      on Press: SetTag("MH_Control_Visibility", 1); SetTag("Press_Control_Screen", 2)
      Visibility <- "DB704_MH_Value_Mixinghead{0}_AmountComponent"
   Button "Button_31" at 489,499 size 94x25; TextOff 'Text'
      on Press: SetTag("MH_Control_Visibility", 2); SetTag("Temp_Control_Screen", 2)
      Visibility <- "DB704_MH_Value_Mixinghead{0}_AmountComponent"
   Button "Button_33" at 489,554 size 94x25; TextOff 'Text'
      on Press: SetTag("MH_Control_Visibility", 2); SetTag("Temp_Control_Screen", 4)
      Visibility <- "DB704_MH_Value_Mixinghead{0}_AmountComponent"
   Button "Button_32" at 489,527 size 94x25; TextOff 'bar'
      on Press: SetTag("MH_Control_Visibility", 1); SetTag("Press_Control_Screen", 4)
      Visibility <- "DB704_MH_Value_Mixinghead{0}_AmountComponent"
   Button "Button_6" at 768,446 size 94x25; TextOff 'Text'
      on Press: SetTag("MH_Control_Visibility", 2); SetTag("Temp_Control_Screen", 1)
      Visibility <- "DB704_MH_Value_Mixinghead{0}_AmountComponent"
   Button "Button_37" at 768,554 size 94x25; TextOff 'Text'
      on Press: SetTag("MH_Control_Visibility", 2); SetTag("Temp_Control_Screen", 5)
      Visibility <- "DB704_MH_Value_Mixinghead{0}_AmountComponent"
   Button "Button_36" at 768,527 size 94x25; TextOff 'bar'
      on Press: SetTag("MH_Control_Visibility", 1); SetTag("Press_Control_Screen", 5)
      Visibility <- "DB704_MH_Value_Mixinghead{0}_AmountComponent"
   Button "Button_35" at 768,499 size 94x25; TextOff 'Text'
      on Press: SetTag("MH_Control_Visibility", 2); SetTag("Temp_Control_Screen", 3)
      Visibility <- "DB704_MH_Value_Mixinghead{0}_AmountComponent"
   Button "Button_34" at 768,473 size 94x25; TextOff 'bar'
      on Press: SetTag("MH_Control_Visibility", 1); SetTag("Press_Control_Screen", 3)
      Visibility <- "DB704_MH_Value_Mixinghead{0}_AmountComponent"
   Button "Button_5" at 768,421 size 94x25; TextOff 'bar'
      on Press: SetTag("MH_Control_Visibility", 1); SetTag("Press_Control_Screen", 1)
      Visibility <- "DB704_MH_Value_Mixinghead{0}_AmountComponent"
   Button "Button_19" at 332,596 size 138x30; TextOff 'Text'; TextList "Pump_Name"
      Visibility <- "DB704_MH_Value_Mixinghead{0}_AmountComponent"
      ProcessValue <- "DB704_MH_Value_Mixinghead{0}_MH_Connection{1}_Pump_No"
      Appearance <- "DB614_MH_State_MH_Connection{0}_colour{1}"
   Button "Button_38" at 470,596 size 138x30; TextOff 'Text'; TextList "Pump_Name"
      Visibility <- "DB704_MH_Value_Mixinghead{0}_AmountComponent"
      ProcessValue <- "DB704_MH_Value_Mixinghead{0}_MH_Connection{2}_Pump_No"
      Appearance <- "DB614_MH_State_MH_Connection{0}_colour{2}"
   Button "Button_40" at 608,596 size 138x30; TextOff 'Text'; TextList "Pump_Name"
      Visibility <- "DB704_MH_Value_Mixinghead{0}_AmountComponent"
      ProcessValue <- "DB704_MH_Value_Mixinghead{0}_MH_Connection{3}_Pump_No"
      Appearance <- "DB614_MH_State_MH_Connection{0}_colour{3}"
   Button "Button_47" at 746,596 size 138x30; TextOff 'Text'; TextList "Pump_Name"
      Visibility <- "DB704_MH_Value_Mixinghead{0}_AmountComponent"
      ProcessValue <- "DB704_MH_Value_Mixinghead{0}_MH_Connection{4}_Pump_No"
      Appearance <- "DB614_MH_State_MH_Connection{0}_colour{4}"
   Button "Button_48" at 884,596 size 138x30; TextOff 'Text'; TextList "Pump_Name"
      Visibility <- "DB704_MH_Value_Mixinghead{0}_AmountComponent"
      ProcessValue <- "DB704_MH_Value_Mixinghead{0}_MH_Connection{5}_Pump_No"
      Appearance <- "DB614_MH_State_MH_Connection{0}_colour{5}"
   Button "Button_49" at 1022,596 size 138x30; TextOff 'Text'; TextList "Pump_Name"
      Visibility <- "DB704_MH_Value_Mixinghead{0}_AmountComponent"
      ProcessValue <- "DB704_MH_Value_Mixinghead{0}_MH_Connection{6}_Pump_No"
      Appearance <- "DB614_MH_State_MH_Connection{0}_colour{6}"
   Button "Button_50" at 342,413 size 138x30; TextOff 'Text'; TextList "Pump_Name"
      Visibility <- "DB704_MH_Value_Mixinghead{0}_AmountComponent"
      ProcessValue <- "DB704_MH_Value_Mixinghead{0}_MH_Connection{1}_Pump_No"
      Appearance <- "DB614_MH_State_MH_Connection{0}_colour{1}"
   Button "Button_51" at 342,474 size 138x30; TextOff 'Text'; TextList "Pump_Name"
      Visibility <- "DB704_MH_Value_Mixinghead{0}_AmountComponent"
      ProcessValue <- "DB704_MH_Value_Mixinghead{0}_MH_Connection{3}_Pump_No"
      Appearance <- "DB614_MH_State_MH_Connection{0}_colour{3}"
   Button "Button_52" at 342,535 size 138x30; TextOff 'Text'; TextList "Pump_Name"
      Visibility <- "DB704_MH_Value_Mixinghead{0}_AmountComponent"
      ProcessValue <- "DB704_MH_Value_Mixinghead{0}_MH_Connection{5}_Pump_No"
      Appearance <- "DB614_MH_State_MH_Connection{0}_colour{5}"
   Button "Button_53" at 871,413 size 138x30; TextOff 'Text'; TextList "Pump_Name"
      Visibility <- "DB704_MH_Value_Mixinghead{0}_AmountComponent"
      ProcessValue <- "DB704_MH_Value_Mixinghead{0}_MH_Connection{2}_Pump_No"
      Appearance <- "DB614_MH_State_MH_Connection{0}_colour{2}"
   Button "Button_54" at 871,474 size 138x30; TextOff 'Text'; TextList "Pump_Name"
      Visibility <- "DB704_MH_Value_Mixinghead{0}_AmountComponent"
      ProcessValue <- "DB704_MH_Value_Mixinghead{0}_MH_Connection{4}_Pump_No"
      Appearance <- "DB614_MH_State_MH_Connection{0}_colour{4}"
   Button "Button_55" at 871,535 size 138x30; TextOff 'Text'; TextList "Pump_Name"
      Visibility <- "DB704_MH_Value_Mixinghead{0}_AmountComponent"
      ProcessValue <- "DB704_MH_Value_Mixinghead{0}_MH_Connection{6}_Pump_No"
      Appearance <- "DB614_MH_State_MH_Connection{0}_colour{6}"
   GraphicView "Graphic view_10" at 600,423 size 40x37; Picture "logoff"
      Visibility <- "DB123_MH_IO_Signals_MH{0}_IN_MH_Prog_No_MH"
   TextField "Text field_54" at 838,273 size 46x25; Text 's'
      Visibility <- "DB704_MH_Value_Mixinghead{0}_Cleaning_Piston_CP_withInterval"
   TextField "Text field_55" at 838,303 size 46x25; Text 's'
      Visibility <- "DB704_MH_Value_Mixinghead{0}_Cleaning_Piston_CP_withInterval"
   TextField "Text field_40" at 202,455 size 94x25; Text 'NL'
      Visibility <- "DB704_MH_Value_Mixinghead{0}_WithInerting"
   TextField "Text field_41" at 202,430 size 94x25; Text 'NL'
      Visibility <- "DB704_MH_Value_Mixinghead{0}_WithInerting"
   Rectangle "Rectangle_11" at 332,627 size 138x40
      Visibility <- "DB614_MH_State_MH_Status{0}_QPB_Values_selected"
   Rectangle "Rectangle_12" at 332,666 size 138x40
      Visibility <- "DB614_MH_State_MH_Status{0}_QPB_Values_selected"
   Rectangle "Rectangle_13" at 332,705 size 138x40
      Visibility <- "DB614_MH_State_MH_Status{0}_QPB_Values_selected"
   Rectangle "Rectangle_14" at 332,744 size 138x40
      Visibility <- "DB614_MH_State_MH_Status{0}_QPB_Values_selected"
   Rectangle "Rectangle_7" at 470,627 size 138x40
      Visibility <- "DB614_MH_State_MH_Status{0}_QPB_Values_selected"
   Rectangle "Rectangle_8" at 470,666 size 138x40
      Visibility <- "DB614_MH_State_MH_Status{0}_QPB_Values_selected"
   Rectangle "Rectangle_9" at 470,705 size 138x40
      Visibility <- "DB614_MH_State_MH_Status{0}_QPB_Values_selected"
   Rectangle "Rectangle_10" at 470,744 size 138x40
      Visibility <- "DB614_MH_State_MH_Status{0}_QPB_Values_selected"
   TextField "Text field_10" at 106,635 size 70x25; Text 'actual:'
   TextField "Text field_11" at 106,673 size 93x25; Text 'Reduced:'
      Visibility <- "DB614_MH_State_MH_Status{0}_QPB_Values_selected"
   TextField "Text field_12" at 106,711 size 144x25; Text 'High pressure:'
      Visibility <- "DB614_MH_State_MH_Status{0}_QPB_Values_selected"
   TextField "Text field_13" at 106,752 size 139x25; Text 'Low pressure:'
      Visibility <- "DB614_MH_State_MH_Status{0}_QPB_Values_selected"
   TextField "Text field_14" at 277,635 size 46x25; Text 'g/s'
   TextField "Text field_16" at 277,673 size 46x25; Text 'g/s'
      Visibility <- "DB614_MH_State_MH_Status{0}_QPB_Values_selected"
   TextField "Text field_17" at 277,711 size 46x25; Text 'g/s'
      Visibility <- "DB614_MH_State_MH_Status{0}_QPB_Values_selected"
   TextField "Text field_18" at 277,749 size 46x25; Text 'bar'
      Visibility <- "DB614_MH_State_MH_Status{0}_QPB_Values_selected"
   Button "reduced icon" at 237,673 size 34x27; TextOff 'Text'; PictureOff "Reduced green"
      Visibility <- "DB614_MH_State_MH_Status{0}_QPB_Values_selected"
   Button "Interval icon" at 237,712 size 34x27; TextOff 'Text'; PictureOff "Interval green"
      Visibility <- "DB614_MH_State_MH_Status{0}_QPB_Values_selected"
   Button "Lowpress icon" at 237,751 size 34x27; TextOff 'Text'; PictureOff "Lowpress green"
      Visibility <- "DB614_MH_State_MH_Status{0}_QPB_Values_selected"
   Rectangle "Rectangle_15" at 608,627 size 138x40
      Visibility <- "DB614_MH_State_MH_Status{0}_QPB_Values_selected"
   Rectangle "Rectangle_16" at 608,666 size 138x40
      Visibility <- "DB614_MH_State_MH_Status{0}_QPB_Values_selected"
   Rectangle "Rectangle_17" at 608,705 size 138x40
      Visibility <- "DB614_MH_State_MH_Status{0}_QPB_Values_selected"
   Rectangle "Rectangle_18" at 608,744 size 138x40
      Visibility <- "DB614_MH_State_MH_Status{0}_QPB_Values_selected"
   Rectangle "Rectangle_19" at 746,627 size 138x40
      Visibility <- "DB614_MH_State_MH_Status{0}_QPB_Values_selected"
   Rectangle "Rectangle_20" at 746,666 size 138x40
      Visibility <- "DB614_MH_State_MH_Status{0}_QPB_Values_selected"
   Rectangle "Rectangle_21" at 746,705 size 138x40
      Visibility <- "DB614_MH_State_MH_Status{0}_QPB_Values_selected"
   Rectangle "Rectangle_22" at 746,744 size 138x40
      Visibility <- "DB614_MH_State_MH_Status{0}_QPB_Values_selected"
   Rectangle "Rectangle_23" at 884,627 size 138x40
      Visibility <- "DB614_MH_State_MH_Status{0}_QPB_Values_selected"
   Rectangle "Rectangle_24" at 884,666 size 138x40
      Visibility <- "DB614_MH_State_MH_Status{0}_QPB_Values_selected"
   Rectangle "Rectangle_25" at 884,705 size 138x40
      Visibility <- "DB614_MH_State_MH_Status{0}_QPB_Values_selected"
   Rectangle "Rectangle_26" at 884,744 size 138x40
      Visibility <- "DB614_MH_State_MH_Status{0}_QPB_Values_selected"
   Rectangle "Rectangle_27" at 1022,627 size 138x40
      Visibility <- "DB614_MH_State_MH_Status{0}_QPB_Values_selected"
   Rectangle "Rectangle_28" at 1022,666 size 138x40
      Visibility <- "DB614_MH_State_MH_Status{0}_QPB_Values_selected"
   Rectangle "Rectangle_29" at 1022,705 size 138x40
      Visibility <- "DB614_MH_State_MH_Status{0}_QPB_Values_selected"
   Rectangle "Rectangle_30" at 1022,744 size 138x40
      Visibility <- "DB614_MH_State_MH_Status{0}_QPB_Values_selected"
   IOField "I/O field_23" at 202,430 size 69x25; FormatPattern 9999.9
      ProcessValue <- "DB614_MH_State_InertingMH{0}_Computed_Value"
      Visibility <- "DB704_MH_Value_Mixinghead{0}_WithInerting"
   IOField "I/O field_24" at 202,455 size 69x25; FormatPattern 9999.9
      ProcessValue <- "DB614_MH_State_InertingMH{0}_Total_Flow_N2_Visu"
      Visibility <- "DB704_MH_Value_Mixinghead{0}_WithInerting"
   Button "b_Reduced_Con1" at 335,670 size 36x32; TextOff 'Text'; PictureList "Check_Uncheck"
      Visibility <- "DB614_MH_State_MH_Status{0}_QPB_Values_selected"
      on Click: InvertBit("DB704_MH_Value_Mixinghead{0}_MH_Connection{1}_Red_CircOverNozzle")
      ProcessValue <- "DB704_MH_Value_Mixinghead{0}_MH_Connection{1}_Red_CircOverNozzle"
   Button "b_HP_Con1" at 335,709 size 36x32; TextOff 'Text'; PictureList "Check_Uncheck"
      Visibility <- "DB614_MH_State_MH_Status{0}_QPB_Values_selected"
      on Click: InvertBit("DB704_MH_Value_Mixinghead{0}_MH_Connection{1}_HP_CircOverNozzle")
      ProcessValue <- "DB704_MH_Value_Mixinghead{0}_MH_Connection{1}_HP_CircOverNozzle"
   Button "b_LP_Con1" at 335,748 size 36x32; TextOff 'Text'; PictureList "Check_Uncheck"
      Visibility <- "DB614_MH_State_MH_Status{0}_QPB_Values_selected"
      on Click: InvertBit("DB704_MH_Value_Mixinghead{0}_MH_Connection{1}_LP_CircOverNozzle")
      ProcessValue <- "DB704_MH_Value_Mixinghead{0}_MH_Connection{1}_LP_CircOverNozzle"
   Button "b_LP_Con2" at 473,748 size 36x32; TextOff 'Text'; PictureList "Check_Uncheck"
      Visibility <- "DB614_MH_State_MH_Status{0}_QPB_Values_selected"
      on Click: InvertBit("DB704_MH_Value_Mixinghead{0}_MH_Connection{2}_LP_CircOverNozzle")
      ProcessValue <- "DB704_MH_Value_Mixinghead{0}_MH_Connection{2}_LP_CircOverNozzle"
   Button "b_HP_Con2" at 473,709 size 36x32; TextOff 'Text'; PictureList "Check_Uncheck"
      Visibility <- "DB614_MH_State_MH_Status{0}_QPB_Values_selected"
      on Click: InvertBit("DB704_MH_Value_Mixinghead{0}_MH_Connection{2}_HP_CircOverNozzle")
      ProcessValue <- "DB704_MH_Value_Mixinghead{0}_MH_Connection{2}_HP_CircOverNozzle"
   Button "b_Reduced_Con2" at 473,670 size 36x32; TextOff 'Text'; PictureList "Check_Uncheck"
      Visibility <- "DB614_MH_State_MH_Status{0}_QPB_Values_selected"
      on Click: InvertBit("DB704_MH_Value_Mixinghead{0}_MH_Connection{2}_Red_CircOverNozzle")
      ProcessValue <- "DB704_MH_Value_Mixinghead{0}_MH_Connection{2}_Red_CircOverNozzle"
   Button "b_Reduced_Con3" at 611,670 size 36x32; TextOff 'Text'; PictureList "Check_Uncheck"
      Visibility <- "DB614_MH_State_MH_Status{0}_QPB_Values_selected"
      on Click: InvertBit("DB704_MH_Value_Mixinghead{0}_MH_Connection{3}_Red_CircOverNozzle")
      ProcessValue <- "DB704_MH_Value_Mixinghead{0}_MH_Connection{3}_Red_CircOverNozzle"
   Button "b_HP_Con3" at 611,709 size 36x32; TextOff 'Text'; PictureList "Check_Uncheck"
      Visibility <- "DB614_MH_State_MH_Status{0}_QPB_Values_selected"
      on Click: InvertBit("DB704_MH_Value_Mixinghead{0}_MH_Connection{3}_HP_CircOverNozzle")
      ProcessValue <- "DB704_MH_Value_Mixinghead{0}_MH_Connection{3}_HP_CircOverNozzle"
   Button "b_LP_Con3" at 611,748 size 36x32; TextOff 'Text'; PictureList "Check_Uncheck"
      Visibility <- "DB614_MH_State_MH_Status{0}_QPB_Values_selected"
      on Click: InvertBit("DB704_MH_Value_Mixinghead{0}_MH_Connection{3}_LP_CircOverNozzle")
      ProcessValue <- "DB704_MH_Value_Mixinghead{0}_MH_Connection{3}_LP_CircOverNozzle"
   Button "b_LP_Con4" at 749,748 size 36x32; TextOff 'Text'; PictureList "Check_Uncheck"
      Visibility <- "DB614_MH_State_MH_Status{0}_QPB_Values_selected"
      on Click: InvertBit("DB704_MH_Value_Mixinghead{0}_MH_Connection{4}_LP_CircOverNozzle")
      ProcessValue <- "DB704_MH_Value_Mixinghead{0}_MH_Connection{4}_LP_CircOverNozzle"
   Button "b_HP_Con4" at 749,709 size 36x32; TextOff 'Text'; PictureList "Check_Uncheck"
      Visibility <- "DB614_MH_State_MH_Status{0}_QPB_Values_selected"
      on Click: InvertBit("DB704_MH_Value_Mixinghead{0}_MH_Connection{4}_HP_CircOverNozzle")
      ProcessValue <- "DB704_MH_Value_Mixinghead{0}_MH_Connection{4}_HP_CircOverNozzle"
   Button "b_Reduced_Con4" at 749,670 size 36x32; TextOff 'Text'; PictureList "Check_Uncheck"
      Visibility <- "DB614_MH_State_MH_Status{0}_QPB_Values_selected"
      on Click: InvertBit("DB704_MH_Value_Mixinghead{0}_MH_Connection{4}_Red_CircOverNozzle")
      ProcessValue <- "DB704_MH_Value_Mixinghead{0}_MH_Connection{4}_Red_CircOverNozzle"
   Button "b_Reduced_Con5" at 887,670 size 36x32; TextOff 'Text'; PictureList "Check_Uncheck"
      Visibility <- "DB614_MH_State_MH_Status{0}_QPB_Values_selected"
      on Click: InvertBit("DB704_MH_Value_Mixinghead{0}_MH_Connection{5}_Red_CircOverNozzle")
      ProcessValue <- "DB704_MH_Value_Mixinghead{0}_MH_Connection{5}_Red_CircOverNozzle"
   Button "b_HP_Con5" at 887,709 size 36x32; TextOff 'Text'; PictureList "Check_Uncheck"
      Visibility <- "DB614_MH_State_MH_Status{0}_QPB_Values_selected"
      on Click: InvertBit("DB704_MH_Value_Mixinghead{0}_MH_Connection{5}_HP_CircOverNozzle")
      ProcessValue <- "DB704_MH_Value_Mixinghead{0}_MH_Connection{5}_HP_CircOverNozzle"
   Button "b_LP_Con5" at 887,748 size 36x32; TextOff 'Text'; PictureList "Check_Uncheck"
      Visibility <- "DB614_MH_State_MH_Status{0}_QPB_Values_selected"
      on Click: InvertBit("DB704_MH_Value_Mixinghead{0}_MH_Connection{5}_LP_CircOverNozzle")
      ProcessValue <- "DB704_MH_Value_Mixinghead{0}_MH_Connection{5}_LP_CircOverNozzle"
   Button "b_LP_Con6" at 1025,748 size 36x32; TextOff 'Text'; PictureList "Check_Uncheck"
      Visibility <- "DB614_MH_State_MH_Status{0}_QPB_Values_selected"
      on Click: InvertBit("DB704_MH_Value_Mixinghead{0}_MH_Connection{6}_LP_CircOverNozzle")
      ProcessValue <- "DB704_MH_Value_Mixinghead{0}_MH_Connection{6}_LP_CircOverNozzle"
   Button "b_HP_Con6" at 1025,709 size 36x32; TextOff 'Text'; PictureList "Check_Uncheck"
      Visibility <- "DB614_MH_State_MH_Status{0}_QPB_Values_selected"
      on Click: InvertBit("DB704_MH_Value_Mixinghead{0}_MH_Connection{6}_HP_CircOverNozzle")
      ProcessValue <- "DB704_MH_Value_Mixinghead{0}_MH_Connection{6}_HP_CircOverNozzle"
   Button "b_Reduced_Con6" at 1025,670 size 36x32; TextOff 'Text'; PictureList "Check_Uncheck"
      Visibility <- "DB614_MH_State_MH_Status{0}_QPB_Values_selected"
      on Click: InvertBit("DB704_MH_Value_Mixinghead{0}_MH_Connection{6}_Red_CircOverNozzle")
      ProcessValue <- "DB704_MH_Value_Mixinghead{0}_MH_Connection{6}_Red_CircOverNozzle"

screen "0010_Pump" 1280x800, template "Navigation"
   on GenerateScreen: SetBit("DB613_Komponent_State_Read"); SetTag("Navigation_7", 2); SetBit("DB608_PV_Metering_Read")
   Button "Button_6" at 120,190 size 375x253; TextOff 'Text'
      Visibility <- "Metering Display Open"
   Button "Button_7" at 443,193 size 51x41; TextOff 'Text'; PictureOff "images (1)"
      on Press: SetTag("NavScreenChange", 0); SetTag("Metering Display Open", 0)
      Visibility <- "Metering Display Open"
   TextField "Text field_4" at 255,213 size 66x29; Text 'Ratio'
      Visibility <- "Metering Display Open"
   TextField "Text field_5" at 133,269 size 72x25; Text 'Actual:'
      Visibility <- "Metering Display Open"
   TextField "Text field_6" at 133,295 size 100x25; Text 'Set value:'
      Visibility <- "Metering Display Open"
   TextField "Text field_7" at 133,319 size 201x25; Text 'Warning upper limit:'
      Visibility <- "Metering Display Open"
   TextField "Text field_8" at 133,345 size 199x25; Text 'Warning lower limit:'
      Visibility <- "Metering Display Open"
   TextField "Text field_9" at 133,371 size 170x25; Text 'Fault upper limit:'
      Visibility <- "Metering Display Open"
   TextField "Text field_10" at 133,397 size 168x25; Text 'Fault lower limit:'
      Visibility <- "Metering Display Open"
   IOField "I/O field_3" at 344,345 size 96x25; Authorization "Operate"; FormatPattern 99.9
      ProcessValue <- "DB608_PV_Metering_Metering{0}_MixingRatio_PV_SetV_WarningLowerLimit"
      Visibility <- "Metering Display Open"
   IOField "I/O field_4" at 344,319 size 96x25; Authorization "Operate"; FormatPattern 99.9
      ProcessValue <- "DB608_PV_Metering_Metering{0}_MixingRatio_PV_SetV_WarningUpperLimit"
      Visibility <- "Metering Display Open"
   IOField "I/O field_6" at 344,397 size 96x25; Authorization "Operate"; FormatPattern 99.9
      ProcessValue <- "DB608_PV_Metering_Metering{0}_MixingRatio_PV_SetV_AlarmLowerLimit"
      Visibility <- "Metering Display Open"
   IOField "I/O field_7" at 344,371 size 96x25; Authorization "Operate"; FormatPattern 99.9
      ProcessValue <- "DB608_PV_Metering_Metering{0}_MixingRatio_PV_SetV_AlarmUpperLimit"
      Visibility <- "Metering Display Open"
   IOField "I/O field_8" at 344,295 size 96x25; FormatPattern 999.9
      ProcessValue <- "DB608_PV_Metering_Metering{0}_MixingRatio_PV_SetV_Value"
      Visibility <- "Metering Display Open"
   IOField "I/O field_9" at 344,269 size 96x25; FormatPattern 999.9
      Visibility <- "Metering Display Open"
      ProcessValue <- "DB608_PV_Metering_Metering{0}_MixingRatio_PV_ActV_Value"
   TextField "Text field_11" at 448,269 size 46x25; Text '%'
      Visibility <- "Metering Display Open"
   TextField "Text field_12" at 448,295 size 46x25; Text '%'
      Visibility <- "Metering Display Open"
   TextField "Text field_13" at 448,321 size 45x25; Text 'Δ %'
      Visibility <- "Metering Display Open"
   TextField "Text field_14" at 448,347 size 45x25; Text 'Δ %'
      Visibility <- "Metering Display Open"
   TextField "Text field_15" at 448,373 size 45x25; Text 'Δ %'
      Visibility <- "Metering Display Open"
   TextField "Text field_16" at 448,399 size 45x25; Text 'Δ %'
      Visibility <- "Metering Display Open"
   Button "Button_2" at 120,190 size 375x253; TextOff 'Text'
      Visibility <- "Metering Display Open"
   Button "Button_4" at 438,194 size 51x41; TextOff 'Text'; PictureOff "images (1)"
      on Press: SetTag("NavScreenChange", 0); SetTag("Metering Display Open", 0)
      Visibility <- "Metering Display Open"
   TextField "Text field_17" at 278,205 size 59x29; Text 'Flow'
      Visibility <- "Metering Display Open"
   TextField "Text field_18" at 133,269 size 72x25; Text 'Actual:'
      Visibility <- "Metering Display Open"
   TextField "Text field_19" at 133,296 size 100x25; Text 'Set value:'
      Visibility <- "Metering Display Open"
   TextField "Text field_20" at 133,320 size 201x25; Text 'Warning upper limit:'
      Visibility <- "Metering Display Open"
   TextField "Text field_21" at 133,347 size 199x25; Text 'Warning lower limit:'
      Visibility <- "Metering Display Open"
   TextField "Text field_22" at 133,373 size 170x25; Text 'Fault upper limit:'
      Visibility <- "Metering Display Open"
   TextField "Text field_23" at 133,400 size 168x25; Text 'Fault lower limit:'
      Visibility <- "Metering Display Open"
   IOField "I/O field_10" at 329,347 size 96x25; Authorization "Operate"; FormatPattern 99.99
      ProcessValue <- "DB608_PV_Metering_Metering{0}_Flow_PV_SetV_WarningLowerLimit"
      Visibility <- "Metering Display Open"
   IOField "I/O field_11" at 329,320 size 96x25; Authorization "Operate"; FormatPattern 99.99
      ProcessValue <- "DB608_PV_Metering_Metering{0}_Flow_PV_SetV_WarningUpperLimit"
      Visibility <- "Metering Display Open"
   IOField "I/O field_12" at 329,400 size 96x25; Authorization "Operate"; FormatPattern 99.99
      ProcessValue <- "DB608_PV_Metering_Metering{0}_Flow_PV_SetV_AlarmLowerLimit"
      Visibility <- "Metering Display Open"
   IOField "I/O field_13" at 329,373 size 96x25; Authorization "Operate"; FormatPattern 99.99
      ProcessValue <- "DB608_PV_Metering_Metering{0}_Flow_PV_SetV_AlarmUpperLimit"
      Visibility <- "Metering Display Open"
   IOField "I/O field_14" at 329,296 size 96x25; FormatPattern 9999.99
      ProcessValue <- "DB608_PV_Metering_Metering{0}_Flow_PV_SetV_Value"
      Visibility <- "Metering Display Open"
   IOField "I/O field_15" at 329,268 size 96x25; FormatPattern 9999.99
      Visibility <- "Metering Display Open"
      ProcessValue <- "DB608_PV_Metering_Metering{0}_Flow_PV_ActV_Value"
   TextField "Text field_24" at 431,269 size 46x25; Text 'g/s'
      Visibility <- "Metering Display Open"
   TextField "Text field_25" at 431,296 size 46x25; Text 'g/s'
      Visibility <- "Metering Display Open"
   TextField "Text field_26" at 431,320 size 57x25; Text 'Δ g/s'
      Visibility <- "Metering Display Open"
   TextField "Text field_27" at 431,347 size 57x25; Text 'Δ g/s'
      Visibility <- "Metering Display Open"
   TextField "Text field_28" at 431,373 size 57x25; Text 'Δ g/s'
      Visibility <- "Metering Display Open"
   TextField "Text field_29" at 431,400 size 57x25; Text 'Δ g/s'
      Visibility <- "Metering Display Open"
   Button "Template_Button_41" at 16,724 size 68x66; TextOff 'Text'; PictureList "Ico_navigation_2"; PictureOff "Setting_Nav_7"; Authorization "User administration"
      on Click: ActivateScreen("0012_Pump Setting", 0)
      ProcessValue <- "Nav_7"
      Visibility <- "NavUserChange"
   Button "Button_5" at 120,190 size 375x253; TextOff 'Text'
      Visibility <- "Metering Display Open"
   Button "Button_8" at 438,194 size 51x41; TextOff 'Text'; PictureOff "images (1)"
      on Press: SetTag("NavScreenChange", 0); SetTag("Metering Display Open", 0)
      Visibility <- "Metering Display Open"
   TextField "Text field_30" at 278,205 size 104x29; Text 'Pressure'
      Visibility <- "Metering Display Open"
   TextField "Text field_31" at 133,269 size 72x25; Text 'Actual:'
      Visibility <- "Metering Display Open"
   TextField "Text field_32" at 133,294 size 100x25; Text 'Set value:'
      Visibility <- "Metering Display Open"
   TextField "Text field_33" at 133,319 size 201x25; Text 'Warning upper limit:'
      Visibility <- "Metering Display Open"
   TextField "Text field_34" at 133,346 size 199x25; Text 'Warning lower limit:'
      Visibility <- "Metering Display Open"
   TextField "Text field_35" at 133,371 size 170x25; Text 'Fault upper limit:'
      Visibility <- "Metering Display Open"
   TextField "Text field_36" at 133,397 size 168x25; Text 'Fault lower limit:'
      Visibility <- "Metering Display Open"
   IOField "I/O field_16" at 336,346 size 96x25; Authorization "Operate"; FormatPattern 999.9
      ProcessValue <- "DB608_PV_Metering_Metering{0}_Pressure_PV_SetV_WarningLowerLimit"
      Visibility <- "Metering Display Open"
   IOField "I/O field_17" at 336,319 size 96x25; Authorization "Operate"; FormatPattern 999.9
      ProcessValue <- "DB608_PV_Metering_Metering{0}_Pressure_PV_SetV_WarningUpperLimit"
      Visibility <- "Metering Display Open"
   IOField "I/O field_18" at 336,397 size 96x25; Authorization "Operate"; FormatPattern 999.9
      ProcessValue <- "DB608_PV_Metering_Metering{0}_Pressure_PV_SetV_AlarmLowerLimit"
      Visibility <- "Metering Display Open"
   IOField "I/O field_19" at 336,371 size 96x25; Authorization "Operate"; FormatPattern 999.9
      ProcessValue <- "DB608_PV_Metering_Metering{0}_Pressure_PV_SetV_AlarmUpperLimit"
      Visibility <- "Metering Display Open"
   IOField "I/O field_20" at 336,294 size 96x25; FormatPattern 999.9
      Visibility <- "Metering Display Open"
      ProcessValue <- "DB608_PV_Metering_Metering{0}_Pressure_PV_SetV_Value"
   IOField "I/O field_21" at 336,269 size 96x25; FormatPattern 999.9
      Visibility <- "Metering Display Open"
      ProcessValue <- "DB608_PV_Metering_Metering{0}_Pressure_PV_ActV_Value"
   TextField "Text field_37" at 436,269 size 46x25; Text 'bar'
      Visibility <- "Metering Display Open"
   TextField "Text field_38" at 436,294 size 46x25; Text 'bar'
      Visibility <- "Metering Display Open"
   TextField "Text field_39" at 436,321 size 55x25; Text 'Δ bar'
      Visibility <- "Metering Display Open"
   TextField "Text field_40" at 436,346 size 55x25; Text 'Δ bar'
      Visibility <- "Metering Display Open"
   TextField "Text field_41" at 436,371 size 55x25; Text 'Δ bar'
      Visibility <- "Metering Display Open"
   TextField "Text field_42" at 436,397 size 55x25; Text 'Δ bar'
      Visibility <- "Metering Display Open"
   Button "Button_13" at 100,190 size 396x253; TextOff 'Text'
      Visibility <- "OpenPidDialog"
   Button "Button_14" at 438,194 size 51x41; TextOff 'Text'; PictureOff "images (1)"
      on Press: SetTag("NavScreenChange", 0); SetTag("OpenPidDialog", 0)
      Visibility <- "OpenPidDialog"
   TextField "Text field_57" at 119,200 size 359x29; Text 'PI (D) Controller feeding pump'
      Visibility <- "OpenPidDialog"
   TextField "Text field_60" at 134,261 size 171x25; Text 'Actual controller:'
      Visibility <- "OpenPidDialog"
   TextField "Text field_61" at 134,289 size 160x25; Text 'Actual pressure:'
      Visibility <- "OpenPidDialog"
   TextField "Text field_62" at 134,316 size 235x25; Text 'Set Pressure FeedPump:'
      Visibility <- "OpenPidDialog"
   TextField "Text field_63" at 134,344 size 181x25; Text 'Proportional term:'
      Visibility <- "OpenPidDialog"
   TextField "Text field_64" at 134,371 size 139x25; Text 'Integral term:'
      Visibility <- "OpenPidDialog"
   TextField "Text field_65" at 134,399 size 159x25; Text 'Derivative term:'
      Visibility <- "OpenPidDialog"
   IOField "I/O field_24" at 358,344 size 96x25; Authorization "Operate"; FormatPattern 999.9
      Visibility <- "OpenPidDialog"
      ProcessValue <- "DB751_auxiliaryDriveMetering_FeedingPumpControler{0}_ProportionalGain"
   IOField "I/O field_25" at 358,316 size 96x25; Authorization "Operate"; FormatPattern 999.9
      Visibility <- "OpenPidDialog"
      ProcessValue <- "DB608_PV_Metering_Metering{0}_Pre_Pressure_PV_SetV_Value"
   IOField "I/O field_26" at 358,399 size 96x25; Authorization "Operate"; FormatPattern 999.9
      Visibility <- "OpenPidDialog"
      ProcessValue <- "DB751_auxiliaryDriveMetering_FeedingPumpControler{0}_DerivativeTime"
   IOField "I/O field_27" at 358,371 size 96x25; Authorization "Operate"; FormatPattern 999.9
      Visibility <- "OpenPidDialog"
      ProcessValue <- "DB751_auxiliaryDriveMetering_FeedingPumpControler{0}_ResetTime"
   IOField "I/O field_28" at 358,289 size 96x25; FormatPattern 999.9
      Visibility <- "OpenPidDialog"
      ProcessValue <- "DB608_PV_Metering_Metering{0}_Pressure_PV_ActV_Value"
   IOField "I/O field_29" at 358,261 size 96x25; FormatPattern 999.9
      Visibility <- "OpenPidDialog"
      ProcessValue <- "DB608_PV_Metering_Metering{0}_Flow_PV_SetV_Value"
   TextField "Text field_66" at 458,261 size 46x25; Text '%'
      Visibility <- "OpenPidDialog"
   TextField "Text field_67" at 458,289 size 46x25; Text 'bar'
      Visibility <- "OpenPidDialog"
   TextField "Text field_68" at 458,316 size 46x25; Text 'bar'
      Visibility <- "OpenPidDialog"
   Button "b_Pump1" at 176,617 size 48x37; TextOff 'Text'
      on Press: ActivateScreen("0024_ActualFaults", 0); SetTag("Alarm_Filter_Tag", 3)
      Visibility <- "DB613_Komponent_State_FeedPump{0}_FLT_Exist"
   Button "b_Pump1_4" at 321,623 size 48x37; TextOff 'Text'
      on Press: ActivateScreen("0024_ActualFaults", 0); SetTag("Alarm_Filter_Tag", 3)
      Visibility <- "DB613_Komponent_State_HeatexchangerLP{0}_Fault_Exist"
   Button "b_Pump1_1" at 515,631 size 48x37; TextOff 'Text'
      on Press: ActivateScreen("0024_ActualFaults", 0); SetTag("Alarm_Filter_Tag", 3)
      Visibility <- "DB613_Komponent_State_EdgeFilter{0}_FLT_Exist"
   Button "b_Pump1_2" at 671,623 size 48x37; TextOff 'Text'
      on Press: ActivateScreen("0024_ActualFaults", 0); SetTag("Alarm_Filter_Tag", 3)
      Visibility <- "DB613_Komponent_State_MeteringPump{0}_FLT_Exist"
   Button "b_Pump1_3" at 858,600 size 48x37; TextOff 'Text'
      on Press: ActivateScreen("0024_ActualFaults", 0); SetTag("Alarm_Filter_Tag", 3)
      Visibility <- "DB613_Komponent_State_HeatexchangerHP{0}_Fault_Exist"
   TextField "Text field_80" at 839,738 size 104x30; Text 'ºC'
      Visibility <- "DB753_MeteringPump_Pump{0}_WithHeating"
   TextField "Text field_59" at 313,735 size 104x30; Text 'ºC'
      Visibility <- "DB753_MeteringPump_Pump{0}_WithLPHeatExchanger"
   TextField "Text field_56" at 176,742 size 107x30; Text '%'
      Visibility <- "DB751_auxiliaryDriveMetering_FeedingPump{0}_Config_With_PresControl"
   TextField "Text field_55" at 176,706 size 107x30; Text 'bar'
      Visibility <- "DB751_auxiliaryDriveMetering_FeedingPump{0}_Config_With_PresControl"
   Button "Button_19" at 636,603 size 145x62; TextOff 'Text'; PictureOff "motor_2"; PictureList "pump"
      ProcessValue <- "DB613_Komponent_State_ReadDeviceNo"
   Button "Button_1" at 507,186 size 485x409; TextOff 'Text'
   TextField "Text field_1" at 640,675 size 140x30; Text 'bar'
   TextField "Text field_2" at 640,713 size 140x30; Text 'g/s'
   TextField "Text field_3" at 640,751 size 140x30; Text '%'
   Button "Button_9" at 634,672 size 152x35; TextOff 'Text'
      on Press: SetTag("Metering Display Open", 1)
   IOField "Pump_Flow" at 640,716 size 97x26; FormatPattern 9999.99
      ProcessValue <- "DB608_PV_Metering_Metering{0}_Flow_PV_ActV_Value"
   IOField "Pump_Level" at 640,754 size 97x26; FormatPattern 9999.9
      ProcessValue <- "DB608_PV_Metering_Metering{0}_MixingRatio_PV_ActV_Value"
   IOField "Pump_Pressure" at 640,678 size 97x26; FormatPattern 9999.9
      ProcessValue <- "DB608_PV_Metering_Metering{0}_Pressure_PV_ActV_Value"
   Button "b_Increase_Pump" at 785,104 size 46x32; TextOff 'Text'; PictureOff "right arrow"
      on Press: function_dd21b452("DB613_Komponent_State_ReadDeviceNo", 1); function_dd21b452("DB612_Tank_State.ReadDeviceNo", 1)
   Button "b_Decress_Pump" at 273,104 size 46x32; TextOff 'Text'; PictureOff "left arrow"
      on Press: function_b9b71300("DB613_Komponent_State_ReadDeviceNo", 1); function_b9b71300("DB612_Tank_State.ReadDeviceNo", 1)
   IOField "I/O field_34" at 313,735 size 78x30; FormatPattern 9999.9
      ProcessValue <- "DB608_PV_Metering_HeatexchangerLP{0}_PV_ActV_Value"
      Visibility <- "DB753_MeteringPump_Pump{0}_WithLPHeatExchanger"
   IOField "I/O field_22" at 176,706 size 78x30; FormatPattern 9999.9
      ProcessValue <- "DB608_PV_Metering_Metering{0}_Pre_Pressure_PV_ActV_Value"
      Visibility <- "DB751_auxiliaryDriveMetering_FeedingPump{0}_Config_With_PresControl"
   IOField "I/O field_23" at 176,742 size 78x30; FormatPattern 9999
      Visibility <- "DB751_auxiliaryDriveMetering_FeedingPump{0}_Config_With_PresControl"
      ProcessValue <- "DB613_Komponent_State_FeedPump{0}_ManipValuePercent"
   Button "Button_15" at 934,362 size 45x30; TextOff 'Text'; PictureOff "obeng"
      on Press: SetTag("OpenPidDialog", 1)
      Visibility <- "DB751_auxiliaryDriveMetering_FeedingPump{0}_Config_With_PresControl"
   TextField "Text field_69" at 896,226 size 46x25; Text 's'
      Visibility <- "DB753_MeteringPump_Pump{0}_WithFeedPump"
   TextField "Text field_70" at 896,253 size 46x25; Text 's'
      Visibility <- "DB753_MeteringPump_Pump{0}_WithFeedPump"
   TextField "Text field_71" at 896,280 size 46x25; Text 's'
      Visibility <- "DB751_auxiliaryDriveMetering_FeedingPump{0}_Config_ManualSwitchON"
   TextField "Text field_72" at 896,308 size 46x25; Text 's'
      Visibility <- "DB751_auxiliaryDriveMetering_FeedingPump{0}_Config_ManualSwitchON"
   TextField "Text field_75" at 896,364 size 46x25; Text 'bar'
      Visibility <- "DB751_auxiliaryDriveMetering_FeedingPump{0}_Config_With_PresControl"
   TextField "Text field_76" at 896,392 size 46x25; Text 's'
      Visibility <- "DB753_MeteringPump_Pump{0}_WithEdgeFilter"
   TextField "Text field_77" at 896,420 size 46x25; Text 's'
      Visibility <- "DB753_MeteringPump_Pump{0}_WithEdgeFilter"
   Button "Button_16" at 933,446 size 45x30; TextOff 'Text'; PictureOff "obeng"
      Visibility <- "DB753_MeteringPump_Pump{0}_WithLPHeatExchanger"
   Button "Button_17" at 933,474 size 45x30; TextOff 'Text'; PictureOff "obeng"
      Visibility <- "DB753_MeteringPump_Pump{0}_WithHeating"
   TextField "Text field_43" at 535,199 size 72x25; Text 'Factor:'
      Visibility <- "DB753_MeteringPump_Pump{0}_WithFlowFactor"
   TextField "Text field_44" at 535,226 size 184x25; Text 'Pre run FeedPump'
      Visibility <- "DB753_MeteringPump_Pump{0}_WithFeedPump"
   TextField "Text field_45" at 535,253 size 217x25; Text 'Delay time FeedPump:'
      Visibility <- "DB753_MeteringPump_Pump{0}_WithFeedPump"
   TextField "Text field_46" at 535,280 size 195x25; Text 'Runtime FeedPump:'
      Visibility <- "DB751_auxiliaryDriveMetering_FeedingPump{0}_Config_ManualSwitchON"
   TextField "Text field_47" at 535,308 size 218x25; Text 'Break time FeedPump:'
      Visibility <- "DB751_auxiliaryDriveMetering_FeedingPump{0}_Config_ManualSwitchON"
   TextField "Text field_48" at 535,336 size 239x25; Text 'Enable temp. FeedPump:'
      Visibility <- "DB753_MeteringPump_Pump{0}_WithMinTempRelease"
   TextField "Text field_49" at 535,364 size 228x25; Text 'Set Pressure FeedPump'
      Visibility <- "DB751_auxiliaryDriveMetering_FeedingPump{0}_Config_With_PresControl"
   TextField "Text field_50" at 535,392 size 193x25; Text 'Runtime EdgeFilter:'
      Visibility <- "DB753_MeteringPump_Pump{0}_WithEdgeFilter"
   TextField "Text field_51" at 535,420 size 211x25; Text 'Pause time EdgeFilter'
      Visibility <- "DB753_MeteringPump_Pump{0}_WithEdgeFilter"
   TextField "Text field_52" at 535,448 size 160x25; Text 'Temp. LP Heater'
      Visibility <- "DB753_MeteringPump_Pump{0}_WithLPHeatExchanger"
   TextField "Text field_53" at 535,476 size 170x25; Text 'Temp. HP Heater:'
      Visibility <- "DB753_MeteringPump_Pump{0}_WithHeating"
   TextField "Text field_54" at 535,558 size 257x25; Text 'Enable temp. comp. pump:'
      Visibility <- "DB753_MeteringPump_Pump{0}_WithMinTempRelease"
   IOField "I/O field_31" at 791,199 size 96x25; Authorization "Operate"; FormatPattern 99999.99
      ProcessValue <- "DB753_MeteringPump_Pump{0}_FlowFactor"
      Visibility <- "DB753_MeteringPump_Pump{0}_WithFlowFactor"
   IOField "I/O field_32" at 791,226 size 96x25; Authorization "Operate"; FormatPattern 99999
      ProcessValue <- "DB753_MeteringPump_Pump{0}_DelayPressureFeedP"
      Visibility <- "DB753_MeteringPump_Pump{0}_WithFeedPump"
   IOField "I/O field_33" at 791,253 size 96x25; Authorization "Operate"; FormatPattern 99999
      ProcessValue <- "DB753_MeteringPump_Pump{0}_DelayRunTimeFeedP"
      Visibility <- "DB753_MeteringPump_Pump{0}_WithFeedPump"
   IOField "I/O field_35" at 791,280 size 96x25; Authorization "Operate"; FormatPattern 99999
      ProcessValue <- "DB751_auxiliaryDriveMetering_FeedingPump{0}_RunTime"
      Visibility <- "DB751_auxiliaryDriveMetering_FeedingPump{0}_Config_ManualSwitchON"
   IOField "I/O field_36" at 791,308 size 96x25; Authorization "Operate"; FormatPattern 99999
      ProcessValue <- "DB751_auxiliaryDriveMetering_FeedingPump{0}_PauseTime"
      Visibility <- "DB751_auxiliaryDriveMetering_FeedingPump{0}_Config_ManualSwitchON"
   IOField "I/O field_37" at 791,336 size 96x25; Authorization "Operate"; FormatPattern 99999
      ProcessValue <- "DB751_auxiliaryDriveMetering_FeedingPump{0}_MinTempRelease"
      Visibility <- "DB753_MeteringPump_Pump{0}_WithMinTempRelease"
   IOField "I/O field_30" at 791,364 size 96x25; Authorization "Operate"; FormatPattern 99999.9
      Visibility <- "DB751_auxiliaryDriveMetering_FeedingPump{0}_Config_With_PresControl"
      ProcessValue <- "DB608_PV_Metering_Metering{0}_Pre_Pressure_PV_SetV_Value"
   IOField "I/O field_38" at 791,392 size 96x25; Authorization "Operate"; FormatPattern 99999
      ProcessValue <- "DB751_auxiliaryDriveMetering_EdgeFilter{0}_RunTime"
      Visibility <- "DB753_MeteringPump_Pump{0}_WithEdgeFilter"
   IOField "I/O field_39" at 791,420 size 96x25; Authorization "Operate"; FormatPattern 99999
      ProcessValue <- "DB751_auxiliaryDriveMetering_EdgeFilter{0}_PauseTime"
      Visibility <- "DB753_MeteringPump_Pump{0}_WithEdgeFilter"
   IOField "I/O field_40" at 791,448 size 96x25; Authorization "Operate"; FormatPattern 99999.9
      ProcessValue <- "DB608_PV_Metering_HeatexchangerLP{0}_PV_SetV_Value"
      Visibility <- "DB753_MeteringPump_Pump{0}_WithLPHeatExchanger"
   IOField "I/O field_41" at 791,476 size 96x25; Authorization "Operate"; FormatPattern 99999.9
      ProcessValue <- "DB608_PV_Metering_HeatexchangerHP{0}_PV_SetV_Value"
      Visibility <- "DB753_MeteringPump_Pump{0}_WithHeating"
   IOField "I/O field_42" at 791,558 size 96x25; Authorization "Operate"; FormatPattern 99999.9
      ProcessValue <- "DB753_MeteringPump_Pump{0}_MinTempRelease"
      Visibility <- "DB753_MeteringPump_Pump{0}_WithMinTempRelease"
   IOField "I/O field_43" at 326,104 size 451x32; Authorization "Operate"; FormatPattern ????????????????????
      ProcessValue <- "DB753_MeteringPump_Pump{0}_Name"
      Appearance <- "DB702_Tank_Value_Tank{0}_Color"
   Button "Button_3" at 1087,208 size 81x116; TextOff 'Text'
      Visibility <- "DB753_MeteringPump_Pump{0}_WithEdgeFilter"
   Rectangle "Rectangle_10" at 1096,218 size 64x56
      Appearance <- "DB613_Komponent_State_EdgeFilter{0}_State_Drive"
      Visibility <- "DB753_MeteringPump_Pump{0}_WithEdgeFilter"
   GraphicIOField "Graphic I/O field_9" at 1104,221 size 48x48; PictureList "ON_OFF_SWITCH"
      ProcessValue <- "DB613_Komponent_State_EdgeFilter{0}_Switch_Drive_ON_OFF"
      Visibility <- "DB753_MeteringPump_Pump{0}_WithEdgeFilter"
   Button "Button_18" at 1000,210 size 81x116; TextOff 'Text'
      Visibility <- "DB751_auxiliaryDriveMetering_FeedingPump{0}_Config_ManualSwitchON"
   GraphicView "Graphic view_8" at 1014,282 size 56x30; Picture "motor"
      Visibility <- "DB751_auxiliaryDriveMetering_FeedingPump{0}_Config_ManualSwitchON"
   Rectangle "Rectangle_11" at 1008,218 size 64x56
      Appearance <- "DB613_Komponent_State_FeedPump{0}_State_Drive"
      Visibility <- "DB751_auxiliaryDriveMetering_FeedingPump{0}_Config_ManualSwitchON"
   GraphicIOField "Graphic I/O field_10" at 1016,221 size 48x48; PictureList "ON_OFF_SWITCH"
      ProcessValue <- "DB613_Komponent_State_FeedPump{0}_Switch_Drive_ON_OFF"
      Visibility <- "DB751_auxiliaryDriveMetering_FeedingPump{0}_Config_ManualSwitchON"
   Button "Button_27" at 996,202 size 88x128; TextOff 'Text'
      on Click: InvertBit("DB613_Komponent_State_FeedPump{0}_Switch_Drive_ON_OFF")
      Visibility <- "DB751_auxiliaryDriveMetering_FeedingPump{0}_Config_ManualSwitchON"
   Button "Button_20" at 1088,338 size 81x116; TextOff 'Text'
      Visibility <- "DB753_MeteringPump_Pump{0}_WithHeating"
   Rectangle "Rectangle_1" at 1097,348 size 64x56
      Appearance <- "DB613_Komponent_State_HeatexchangerHP{0}_State_Temp"
      Visibility <- "DB753_MeteringPump_Pump{0}_WithHeating"
   GraphicIOField "Graphic I/O field_1" at 1105,351 size 48x48; PictureList "ON_OFF_SWITCH"
      ProcessValue <- "DB613_Komponent_State_HeatexchangerHP{0}_Switch_Temp_ON_OFF"
      Visibility <- "DB753_MeteringPump_Pump{0}_WithHeating"
   Button "Button_21" at 1000,339 size 81x116; TextOff 'Text'
      Visibility <- "DB753_MeteringPump_Pump{0}_WithLPHeatExchanger"
   Rectangle "Rectangle_3" at 1009,349 size 64x56
      Appearance <- "DB613_Komponent_State_HeatexchangerLP{0}_State_Temp"
      Visibility <- "DB753_MeteringPump_Pump{0}_WithLPHeatExchanger"
   GraphicIOField "Graphic I/O field_2" at 1017,352 size 48x48; PictureList "ON_OFF_SWITCH"
      ProcessValue <- "DB613_Komponent_State_HeatexchangerLP{0}_Switch_Temp_ON_OFF"
      Visibility <- "DB753_MeteringPump_Pump{0}_WithLPHeatExchanger"
   IOField "I/O field_1" at 839,738 size 78x30; FormatPattern 9999.9
      ProcessValue <- "DB608_PV_Metering_HeatexchangerHP{0}_PV_ActV_Value"
      Visibility <- "DB753_MeteringPump_Pump{0}_WithHeating"
   GraphicView "Graphic view_1" at 186,654 size 81x40; Picture "motor2"
      Visibility <- "DB753_MeteringPump_Pump{0}_WithFeedPump"
   GraphicView "Graphic view_2" at 188,627 size 25x21; Picture "AlarmState2"
      Visibility <- "DB613_Komponent_State_FeedPump{0}_FLT_Exist"
   GraphicView "Graphic view_3" at 827,618 size 125x120; Picture "heatHP"
      Visibility <- "DB753_MeteringPump_Pump{0}_WithHeating"
   GraphicView "Graphic view_4" at 871,608 size 25x21; Picture "AlarmState2"
      Visibility <- "DB613_Komponent_State_HeatexchangerHP{0}_Fault_Exist"
   GraphicView "Graphic view_7" at 506,650 size 67x93; Picture "edgefilter"
      Visibility <- "DB753_MeteringPump_Pump{0}_WithEdgeFilter"
   GraphicView "Graphic view_5" at 315,633 size 58x89; Picture "heatLP"
      Visibility <- "DB753_MeteringPump_Pump{0}_WithLPHeatExchanger"
   GraphicView "Graphic view_9" at 380,645 size 39x75; Picture "Graphic_14"
      Visibility <- "DB753_MeteringPump_Pump{0}_WithFischerValveLP"
   GraphicView "Graphic view_10" at 912,639 size 39x75; Picture "Graphic_14"
      Visibility <- "DB753_MeteringPump_Pump{0}_WithFischerValveHP"
   GraphicView "Graphic view_15" at 1003,410 size 76x43; Picture "Switch heatLP"
      Visibility <- "DB753_MeteringPump_Pump{0}_WithLPHeatExchanger"
   Button "Button_24" at 997,333 size 88x128; TextOff 'Text'
      on Click: InvertBit("DB613_Komponent_State_HeatexchangerLP{0}_Switch_Temp_ON_OFF")
      Visibility <- "DB753_MeteringPump_Pump{0}_WithLPHeatExchanger"
   GraphicView "Graphic view_11" at 1105,275 size 44x43; Picture "edgefilter"
      Visibility <- "DB753_MeteringPump_Pump{0}_WithEdgeFilter"
   Button "Button_26" at 1084,202 size 88x128; TextOff 'Text'
      on Click: InvertBit("DB613_Komponent_State_EdgeFilter{0}_Switch_Drive_ON_OFF")
      Visibility <- "DB753_MeteringPump_Pump{0}_WithEdgeFilter"
   GraphicView "Graphic view_14" at 1087,406 size 79x52; Picture "SWITCH HEATHP"
      Visibility <- "DB753_MeteringPump_Pump{0}_WithHeating"
   Button "Button_23" at 1085,332 size 88x128; TextOff 'Text'
      on Click: InvertBit("DB613_Komponent_State_HeatexchangerHP{0}_Switch_Temp_ON_OFF")
      Visibility <- "DB753_MeteringPump_Pump{0}_WithHeating"
   GraphicView "Graphic view_6" at 526,639 size 25x21; Picture "AlarmState2"
      Visibility <- "DB613_Komponent_State_EdgeFilter{0}_FLT_Exist"
   GraphicView "Graphic view_12" at 680,629 size 25x21; Picture "AlarmState2"
      Visibility <- "DB613_Komponent_State_MeteringPump{0}_FLT_Exist"
   GraphicView "Graphic view_13" at 334,631 size 25x21; Picture "AlarmState2"
      Visibility <- "DB613_Komponent_State_HeatexchangerLP{0}_Fault_Exist"
   TextField "Text field_73" at 896,336 size 46x25; Text 'ºC'
      Visibility <- "DB753_MeteringPump_Pump{0}_WithMinTempRelease"
   TextField "Text field_74" at 896,448 size 46x25; Text 'ºC'
      Visibility <- "DB753_MeteringPump_Pump{0}_WithLPHeatExchanger"
   TextField "Text field_78" at 896,558 size 46x25; Text 'ºC'
      Visibility <- "DB753_MeteringPump_Pump{0}_WithMinTempRelease"
   TextField "Text field_79" at 896,476 size 46x25; Text 'ºC'
      Visibility <- "DB753_MeteringPump_Pump{0}_WithHeating"
   Button "Button_12" at 633,673 size 152x35; TextOff 'Text'
      on Press: SetTag("Metering Display Open", 1)
   Button "Button_10" at 633,710 size 152x35; TextOff 'Text'
      on Press: SetTag("Metering Display Open", 2)
   Button "Button_11" at 633,748 size 152x35; TextOff 'Text'
      on Press: SetTag("Metering Display Open", 3)

